      on ChangeValue: SetBit("DB704_MH_Value_Write")
   "DB604_PV_Mixinghead_Mixinghead{0}_Temperature_Connection{2}_PV_Conf_ActV_MaxValueSensor" : Real = PLC DB604_PV_Mixinghead.Mixinghead[0].Temperature_Connection[2].PV_Conf_ActV.MaxValueSensor AT %DB604.DBD382, 1 s
      on ChangeValue: SetBit("DB704_MH_Value_Write")
   "DB604_PV_Mixinghead_Mixinghead{0}_Temperature_Connection{2}_PV_Conf_ActV_MaxSignalResolution" : Real = PLC DB604_PV_Mixinghead.Mixinghead[0].Temperature_Connection[2].PV_Conf_ActV.MaxSignalResolution AT %DB604.DBD386, 1 s
      on ChangeValue: SetBit("DB704_MH_Value_Write")
   "DB604_PV_Mixinghead_Mixinghead{0}_Temperature_Connection{3}_PV_Conf_ActV_ModulNo" : Int = PLC DB604_PV_Mixinghead.Mixinghead[0].Temperature_Connection[3].PV_Conf_ActV.ModulNo AT %DB604.DBW416, 1 s
      on ChangeValue: SetBit("DB704_MH_Value_Write")
   "DB604_PV_Mixinghead_Mixinghead{0}_Temperature_Connection{3}_PV_Conf_ActV_Address" : Int = PLC DB604_PV_Mixinghead.Mixinghead[0].Temperature_Connection[3].PV_Conf_ActV.Address AT %DB604.DBW418, 1 s
      on ChangeValue: SetBit("DB704_MH_Value_Write")
   "DB604_PV_Mixinghead_Mixinghead{0}_Temperature_Connection{3}_PV_Conf_ActV_OffsetSignal" : Int = PLC DB604_PV_Mixinghead.Mixinghead[0].Temperature_Connection[3].PV_Conf_ActV.OffsetSignal AT %DB604.DBW420, 1 s
      on ChangeValue: SetBit("DB704_MH_Value_Write")
   "DB604_PV_Mixinghead_Mixinghead{0}_Temperature_Connection{3}_PV_Conf_ActV_Multiplier" : Real = PLC DB604_PV_Mixinghead.Mixinghead[0].Temperature_Connection[3].PV_Conf_ActV.Multiplier AT %DB604.DBD422, 1 s
      on ChangeValue: SetBit("DB704_MH_Value_Write")
   "DB604_PV_Mixinghead_Mixinghead{0}_Temperature_Connection{3}_PV_Conf_ActV_MinValueSensor" : Real = PLC DB604_PV_Mixinghead.Mixinghead[0].Temperature_Connection[3].PV_Conf_ActV.MinValueSensor AT %DB604.DBD426, 1 s
      on ChangeValue: SetBit("DB704_MH_Value_Write")
   "DB604_PV_Mixinghead_Mixinghead{0}_Temperature_Connection{3}_PV_Conf_ActV_MaxValueSensor" : Real = PLC DB604_PV_Mixinghead.Mixinghead[0].Temperature_Connection[3].PV_Conf_ActV.MaxValueSensor AT %DB604.DBD430, 1 s
      on ChangeValue: SetBit("DB704_MH_Value_Write")
   "DB604_PV_Mixinghead_Mixinghead{0}_Temperature_Connection{3}_PV_Conf_ActV_MaxSignalResolution" : Real = PLC DB604_PV_Mixinghead.Mixinghead[0].Temperature_Connection[3].PV_Conf_ActV.MaxSignalResolution AT %DB604.DBD434, 1 s
      on ChangeValue: SetBit("DB704_MH_Value_Write")
   "DB604_PV_Mixinghead_Mixinghead{0}_Temperature_Connection{4}_PV_Conf_ActV_ModulNo" : Int = PLC DB604_PV_Mixinghead.Mixinghead[0].Temperature_Connection[4].PV_Conf_ActV.ModulNo AT %DB604.DBW464, 1 s
      on ChangeValue: SetBit("DB704_MH_Value_Write")
   "DB604_PV_Mixinghead_Mixinghead{0}_Temperature_Connection{4}_PV_Conf_ActV_Address" : Int = PLC DB604_PV_Mixinghead.Mixinghead[0].Temperature_Connection[4].PV_Conf_ActV.Address AT %DB604.DBW466, 1 s
      on ChangeValue: SetBit("DB704_MH_Value_Write")
   "DB604_PV_Mixinghead_Mixinghead{0}_Temperature_Connection{4}_PV_Conf_ActV_OffsetSignal" : Int = PLC DB604_PV_Mixinghead.Mixinghead[0].Temperature_Connection[4].PV_Conf_ActV.OffsetSignal AT %DB604.DBW468, 1 s
      on ChangeValue: SetBit("DB704_MH_Value_Write")
   "DB604_PV_Mixinghead_Mixinghead{0}_Temperature_Connection{4}_PV_Conf_ActV_Multiplier" : Real = PLC DB604_PV_Mixinghead.Mixinghead[0].Temperature_Connection[4].PV_Conf_ActV.Multiplier AT %DB604.DBD470, 1 s
      on ChangeValue: SetBit("DB704_MH_Value_Write")
   "DB604_PV_Mixinghead_Mixinghead{0}_Temperature_Connection{4}_PV_Conf_ActV_MinValueSensor" : Real = PLC DB604_PV_Mixinghead.Mixinghead[0].Temperature_Connection[4].PV_Conf_ActV.MinValueSensor AT %DB604.DBD474, 1 s
      on ChangeValue: SetBit("DB704_MH_Value_Write")
   "DB604_PV_Mixinghead_Mixinghead{0}_Temperature_Connection{4}_PV_Conf_ActV_MaxValueSensor" : Real = PLC DB604_PV_Mixinghead.Mixinghead[0].Temperature_Connection[4].PV_Conf_ActV.MaxValueSensor AT %DB604.DBD478, 1 s
      on ChangeValue: SetBit("DB704_MH_Value_Write")
   "DB604_PV_Mixinghead_Mixinghead{0}_Temperature_Connection{4}_PV_Conf_ActV_MaxSignalResolution" : Real = PLC DB604_PV_Mixinghead.Mixinghead[0].Temperature_Connection[4].PV_Conf_ActV.MaxSignalResolution AT %DB604.DBD482, 1 s
      on ChangeValue: SetBit("DB704_MH_Value_Write")
   "DB604_PV_Mixinghead_Mixinghead{0}_Temperature_Connection{5}_PV_Conf_ActV_ModulNo" : Int = PLC DB604_PV_Mixinghead.Mixinghead[0].Temperature_Connection[5].PV_Conf_ActV.ModulNo AT %DB604.DBW512, 1 s
      on ChangeValue: SetBit("DB704_MH_Value_Write")
   "DB604_PV_Mixinghead_Mixinghead{0}_Temperature_Connection{5}_PV_Conf_ActV_Address" : Int = PLC DB604_PV_Mixinghead.Mixinghead[0].Temperature_Connection[5].PV_Conf_ActV.Address AT %DB604.DBW514, 1 s
      on ChangeValue: SetBit("DB704_MH_Value_Write")
   "DB604_PV_Mixinghead_Mixinghead{0}_Temperature_Connection{5}_PV_Conf_ActV_OffsetSignal" : Int = PLC DB604_PV_Mixinghead.Mixinghead[0].Temperature_Connection[5].PV_Conf_ActV.OffsetSignal AT %DB604.DBW516, 1 s
      on ChangeValue: SetBit("DB704_MH_Value_Write")
   "DB604_PV_Mixinghead_Mixinghead{0}_Temperature_Connection{5}_PV_Conf_ActV_Multiplier" : Real = PLC DB604_PV_Mixinghead.Mixinghead[0].Temperature_Connection[5].PV_Conf_ActV.Multiplier AT %DB604.DBD518, 1 s
      on ChangeValue: SetBit("DB704_MH_Value_Write")
   "DB604_PV_Mixinghead_Mixinghead{0}_Temperature_Connection{5}_PV_Conf_ActV_MinValueSensor" : Real = PLC DB604_PV_Mixinghead.Mixinghead[0].Temperature_Connection[5].PV_Conf_ActV.MinValueSensor AT %DB604.DBD522, 1 s
      on ChangeValue: SetBit("DB704_MH_Value_Write")
   "DB604_PV_Mixinghead_Mixinghead{0}_Temperature_Connection{5}_PV_Conf_ActV_MaxValueSensor" : Real = PLC DB604_PV_Mixinghead.Mixinghead[0].Temperature_Connection[5].PV_Conf_ActV.MaxValueSensor AT %DB604.DBD526, 1 s
      on ChangeValue: SetBit("DB704_MH_Value_Write")
   "DB604_PV_Mixinghead_Mixinghead{0}_Temperature_Connection{5}_PV_Conf_ActV_MaxSignalResolution" : Real = PLC DB604_PV_Mixinghead.Mixinghead[0].Temperature_Connection[5].PV_Conf_ActV.MaxSignalResolution AT %DB604.DBD530, 1 s
      on ChangeValue: SetBit("DB704_MH_Value_Write")
   "DB604_PV_Mixinghead_Mixinghead{0}_Temperature_Connection{6}_PV_Conf_ActV_ModulNo" : Int = PLC DB604_PV_Mixinghead.Mixinghead[0].Temperature_Connection[6].PV_Conf_ActV.ModulNo AT %DB604.DBW560, 1 s
      on ChangeValue: SetBit("DB704_MH_Value_Write")
   "DB604_PV_Mixinghead_Mixinghead{0}_Temperature_Connection{6}_PV_Conf_ActV_Address" : Int = PLC DB604_PV_Mixinghead.Mixinghead[0].Temperature_Connection[6].PV_Conf_ActV.Address AT %DB604.DBW562, 1 s
      on ChangeValue: SetBit("DB704_MH_Value_Write")
   "DB604_PV_Mixinghead_Mixinghead{0}_Temperature_Connection{6}_PV_Conf_ActV_OffsetSignal" : Int = PLC DB604_PV_Mixinghead.Mixinghead[0].Temperature_Connection[6].PV_Conf_ActV.OffsetSignal AT %DB604.DBW564, 1 s
      on ChangeValue: SetBit("DB704_MH_Value_Write")
   "DB604_PV_Mixinghead_Mixinghead{0}_Temperature_Connection{6}_PV_Conf_ActV_Multiplier" : Real = PLC DB604_PV_Mixinghead.Mixinghead[0].Temperature_Connection[6].PV_Conf_ActV.Multiplier AT %DB604.DBD566, 1 s
      on ChangeValue: SetBit("DB704_MH_Value_Write")
   "DB604_PV_Mixinghead_Mixinghead{0}_Temperature_Connection{6}_PV_Conf_ActV_MinValueSensor" : Real = PLC DB604_PV_Mixinghead.Mixinghead[0].Temperature_Connection[6].PV_Conf_ActV.MinValueSensor AT %DB604.DBD570, 1 s
      on ChangeValue: SetBit("DB704_MH_Value_Write")
   "DB604_PV_Mixinghead_Mixinghead{0}_Temperature_Connection{6}_PV_Conf_ActV_MaxValueSensor" : Real = PLC DB604_PV_Mixinghead.Mixinghead[0].Temperature_Connection[6].PV_Conf_ActV.MaxValueSensor AT %DB604.DBD574, 1 s
      on ChangeValue: SetBit("DB704_MH_Value_Write")
   "DB604_PV_Mixinghead_Mixinghead{0}_Temperature_Connection{6}_PV_Conf_ActV_MaxSignalResolution" : Real = PLC DB604_PV_Mixinghead.Mixinghead[0].Temperature_Connection[6].PV_Conf_ActV.MaxSignalResolution AT %DB604.DBD578, 1 s
      on ChangeValue: SetBit("DB704_MH_Value_Write")
   "DB608_PV_Metering_Metering{0}_MixingRatio_PV_ActV_Value" : Real = PLC DB608_PV_Metering.Metering[0].MixingRatio.PV_ActV.Value AT %DB608.DBD218, 1 s
   "DB608_PV_Metering_HeatexchangerLP{0}_PV_ActV_Value" : Real = PLC DB608_PV_Metering.HeatexchangerLP[0].PV_ActV.Value AT %DB608.DBD3770, 1 s

HMI tags "Last Shot"
   "DB918_ShotResultlast10_FilteredShot{1}_MHNo" : Byte = PLC DB918_ShotResultlast10.FilteredShot[1].MHNo AT %DB918.DBB20, 1 s
   "DB918_ShotResultlast10_FilteredShot{1}_FoamingTime" : Real = PLC DB918_ShotResultlast10.FilteredShot[1].FoamingTime AT %DB918.DBD6, 1 s
   "DB918_ShotResultlast10_FilteredShot{1}_PartWeight" : Real = PLC DB918_ShotResultlast10.FilteredShot[1].PartWeight AT %DB918.DBD10, 1 s
   "DB918_ShotResultlast10_FilteredShot{1}_StationNo" : Byte = PLC DB918_ShotResultlast10.FilteredShot[1].StationNo AT %DB918.DBB18, 1 s
   "DB918_ShotResultlast10_FilteredShot{1}_PartNo" : Int = PLC DB918_ShotResultlast10.FilteredShot[1].PartNo AT %DB918.DBW2, 1 s
   "DB918_ShotResultlast10_FilteredShot{1}_Name{1}" : String[20] = PLC DB918_ShotResultlast10.FilteredShot[1].Name[1] AT %DB918.DBX22.0, 1 s
   "DB918_ShotResultlast10_FilteredShot{1}_Name{2}" : String[20] = PLC DB918_ShotResultlast10.FilteredShot[1].Name[2] AT %DB918.DBX44.0, 1 s
   "DB918_ShotResultlast10_FilteredShot{1}_Flow{1}" : Real = PLC DB918_ShotResultlast10.FilteredShot[1].Flow[1] AT %DB918.DBD154, 1 s
   "DB918_ShotResultlast10_FilteredShot{1}_Flow{2}" : Real = PLC DB918_ShotResultlast10.FilteredShot[1].Flow[2] AT %DB918.DBD158, 1 s
   "DB918_ShotResultlast10_FilteredShot{1}_Pressure{1}" : Real = PLC DB918_ShotResultlast10.FilteredShot[1].Pressure[1] AT %DB918.DBD178, 1 s
   "DB918_ShotResultlast10_FilteredShot{1}_Pressure{2}" : Real = PLC DB918_ShotResultlast10.FilteredShot[1].Pressure[2] AT %DB918.DBD182, 1 s
   "DB918_ShotResultlast10_FilteredShot{1}_Temperature{1}" : Real = PLC DB918_ShotResultlast10.FilteredShot[1].Temperature[1] AT %DB918.DBD202, 1 s
   "DB918_ShotResultlast10_FilteredShot{1}_Temperature{2}" : Real = PLC DB918_ShotResultlast10.FilteredShot[1].Temperature[2] AT %DB918.DBD206, 1 s
   "DB918_ShotResultlast10_FilteredShot{1}_Mixingratio{1}" : Real = PLC DB918_ShotResultlast10.FilteredShot[1].Mixingratio[1] AT %DB918.DBD250, 1 s
   "DB918_ShotResultlast10_FilteredShot{1}_Mixingratio{2}" : Real = PLC DB918_ShotResultlast10.FilteredShot[1].Mixingratio[2] AT %DB918.DBD254, 1 s
   "DB918_ShotResultlast10_FilteredShot{1}_MaterialConsumption{1}" : Real = PLC DB918_ShotResultlast10.FilteredShot[1].MaterialConsumption[1] AT %DB918.DBD226, 1 s
   "DB918_ShotResultlast10_FilteredShot{1}_MaterialConsumption{2}" : Real = PLC DB918_ShotResultlast10.FilteredShot[1].MaterialConsumption[2] AT %DB918.DBD230, 1 s
   "DB918_ShotResultlast10_FilteredShot{2}_PartNo" : Int = PLC DB918_ShotResultlast10.FilteredShot[2].PartNo AT %DB918.DBW288, 1 s
   "DB918_ShotResultlast10_FilteredShot{2}_FoamingTime" : Real = PLC DB918_ShotResultlast10.FilteredShot[2].FoamingTime AT %DB918.DBD292, 1 s
   "DB918_ShotResultlast10_FilteredShot{2}_PartWeight" : Real = PLC DB918_ShotResultlast10.FilteredShot[2].PartWeight AT %DB918.DBD296, 1 s
   "DB918_ShotResultlast10_FilteredShot{2}_StationNo" : Byte = PLC DB918_ShotResultlast10.FilteredShot[2].StationNo AT %DB918.DBB304, 1 s
   "DB918_ShotResultlast10_FilteredShot{2}_MHNo" : Byte = PLC DB918_ShotResultlast10.FilteredShot[2].MHNo AT %DB918.DBB306, 1 s
   "DB918_ShotResultlast10_FilteredShot{2}_Name{1}" : String[20] = PLC DB918_ShotResultlast10.FilteredShot[2].Name[1] AT %DB918.DBX308.0, 1 s
   "DB918_ShotResultlast10_FilteredShot{2}_Name{2}" : String[20] = PLC DB918_ShotResultlast10.FilteredShot[2].Name[2] AT %DB918.DBX330.0, 1 s
   "DB918_ShotResultlast10_FilteredShot{2}_Flow{1}" : Real = PLC DB918_ShotResultlast10.FilteredShot[2].Flow[1] AT %DB918.DBD440, 1 s
   "DB918_ShotResultlast10_FilteredShot{2}_Flow{2}(1)" : Real = PLC DB918_ShotResultlast10.FilteredShot[2].Flow[2] AT %DB918.DBD444, 1 s
   "DB918_ShotResultlast10_FilteredShot{2}_Pressure{1}" : Real = PLC DB918_ShotResultlast10.FilteredShot[2].Pressure[1] AT %DB918.DBD464, 1 s
   "DB918_ShotResultlast10_FilteredShot{2}_Pressure{2}" : Real = PLC DB918_ShotResultlast10.FilteredShot[2].Pressure[2] AT %DB918.DBD468, 1 s
   "DB918_ShotResultlast10_FilteredShot{2}_Temperature{1}" : Real = PLC DB918_ShotResultlast10.FilteredShot[2].Temperature[1] AT %DB918.DBD488, 1 s
   "DB918_ShotResultlast10_FilteredShot{2}_Temperature{2}" : Real = PLC DB918_ShotResultlast10.FilteredShot[2].Temperature[2] AT %DB918.DBD492, 1 s
   "DB918_ShotResultlast10_FilteredShot{2}_MaterialConsumption{1}" : Real = PLC DB918_ShotResultlast10.FilteredShot[2].MaterialConsumption[1] AT %DB918.DBD512, 1 s
   "DB918_ShotResultlast10_FilteredShot{2}_MaterialConsumption{2}" : Real = PLC DB918_ShotResultlast10.FilteredShot[2].MaterialConsumption[2] AT %DB918.DBD516, 1 s
   "DB918_ShotResultlast10_FilteredShot{2}_Mixingratio{1}" : Real = PLC DB918_ShotResultlast10.FilteredShot[2].Mixingratio[1] AT %DB918.DBD536, 1 s
   "DB918_ShotResultlast10_FilteredShot{2}_Mixingratio{2}" : Real = PLC DB918_ShotResultlast10.FilteredShot[2].Mixingratio[2] AT %DB918.DBD540, 1 s
   "DB918_ShotResultlast10_FilteredShot{3}_PartNo" : Int = PLC DB918_ShotResultlast10.FilteredShot[3].PartNo AT %DB918.DBW574, 1 s
   "DB918_ShotResultlast10_FilteredShot{3}_FoamingTime" : Real = PLC DB918_ShotResultlast10.FilteredShot[3].FoamingTime AT %DB918.DBD578, 1 s
   "DB918_ShotResultlast10_FilteredShot{3}_PartWeight" : Real = PLC DB918_ShotResultlast10.FilteredShot[3].PartWeight AT %DB918.DBD582, 1 s
   "DB918_ShotResultlast10_FilteredShot{3}_StationNo" : Byte = PLC DB918_ShotResultlast10.FilteredShot[3].StationNo AT %DB918.DBB590, 1 s
   "DB918_ShotResultlast10_FilteredShot{3}_MHNo" : Byte = PLC DB918_ShotResultlast10.FilteredShot[3].MHNo AT %DB918.DBB592, 1 s
   "DB918_ShotResultlast10_FilteredShot{3}_Name{1}" : String[20] = PLC DB918_ShotResultlast10.FilteredShot[3].Name[1] AT %DB918.DBX594.0, 1 s
   "DB918_ShotResultlast10_FilteredShot{3}_Name{2}" : String[20] = PLC DB918_ShotResultlast10.FilteredShot[3].Name[2] AT %DB918.DBX616.0, 1 s
   "DB918_ShotResultlast10_FilteredShot{3}_Flow{1}" : Real = PLC DB918_ShotResultlast10.FilteredShot[3].Flow[1] AT %DB918.DBD726, 1 s
   "DB918_ShotResultlast10_FilteredShot{3}_Flow{2}" : Real = PLC DB918_ShotResultlast10.FilteredShot[3].Flow[2] AT %DB918.DBD730, 1 s
   "DB918_ShotResultlast10_FilteredShot{3}_Pressure{1}" : Real = PLC DB918_ShotResultlast10.FilteredShot[3].Pressure[1] AT %DB918.DBD750, 1 s
   "DB918_ShotResultlast10_FilteredShot{3}_Pressure{2}" : Real = PLC DB918_ShotResultlast10.FilteredShot[3].Pressure[2] AT %DB918.DBD754, 1 s
   "DB918_ShotResultlast10_FilteredShot{3}_Temperature{1}" : Real = PLC DB918_ShotResultlast10.FilteredShot[3].Temperature[1] AT %DB918.DBD774, 1 s
   "DB918_ShotResultlast10_FilteredShot{3}_Temperature{2}" : Real = PLC DB918_ShotResultlast10.FilteredShot[3].Temperature[2] AT %DB918.DBD778, 1 s
   "DB918_ShotResultlast10_FilteredShot{3}_MaterialConsumption{1}" : Real = PLC DB918_ShotResultlast10.FilteredShot[3].MaterialConsumption[1] AT %DB918.DBD798, 1 s
   "DB918_ShotResultlast10_FilteredShot{3}_MaterialConsumption{2}" : Real = PLC DB918_ShotResultlast10.FilteredShot[3].MaterialConsumption[2] AT %DB918.DBD802, 1 s
   "DB918_ShotResultlast10_FilteredShot{3}_Mixingratio{1}" : Real = PLC DB918_ShotResultlast10.FilteredShot[3].Mixingratio[1] AT %DB918.DBD822, 1 s
   "DB918_ShotResultlast10_FilteredShot{3}_Mixingratio{2}" : Real = PLC DB918_ShotResultlast10.FilteredShot[3].Mixingratio[2] AT %DB918.DBD826, 1 s
   "DB918_ShotResultlast10_FilteredShot{4}_PartNo" : Int = PLC DB918_ShotResultlast10.FilteredShot[4].PartNo AT %DB918.DBW860, 1 s
   "DB918_ShotResultlast10_FilteredShot{4}_FoamingTime" : Real = PLC DB918_ShotResultlast10.FilteredShot[4].FoamingTime AT %DB918.DBD864, 1 s
   "DB918_ShotResultlast10_FilteredShot{4}_PartWeight" : Real = PLC DB918_ShotResultlast10.FilteredShot[4].PartWeight AT %DB918.DBD868, 1 s
   "DB918_ShotResultlast10_FilteredShot{4}_StationNo" : Byte = PLC DB918_ShotResultlast10.FilteredShot[4].StationNo AT %DB918.DBB876, 1 s
   "DB918_ShotResultlast10_FilteredShot{4}_MHNo" : Byte = PLC DB918_ShotResultlast10.FilteredShot[4].MHNo AT %DB918.DBB878, 1 s
   "DB918_ShotResultlast10_FilteredShot{4}_Name{1}" : String[20] = PLC DB918_ShotResultlast10.FilteredShot[4].Name[1] AT %DB918.DBX880.0, 1 s
   "DB918_ShotResultlast10_FilteredShot{4}_Name{2}" : String[20] = PLC DB918_ShotResultlast10.FilteredShot[4].Name[2] AT %DB918.DBX902.0, 1 s
   "DB918_ShotResultlast10_FilteredShot{4}_Flow{1}" : Real = PLC DB918_ShotResultlast10.FilteredShot[4].Flow[1] AT %DB918.DBD1012, 1 s
   "DB918_ShotResultlast10_FilteredShot{4}_Flow{2}" : Real = PLC DB918_ShotResultlast10.FilteredShot[4].Flow[2] AT %DB918.DBD1016, 1 s
   "DB918_ShotResultlast10_FilteredShot{4}_Pressure{1}" : Real = PLC DB918_ShotResultlast10.FilteredShot[4].Pressure[1] AT %DB918.DBD1036, 1 s
   "DB918_ShotResultlast10_FilteredShot{4}_Pressure{2}" : Real = PLC DB918_ShotResultlast10.FilteredShot[4].Pressure[2] AT %DB918.DBD1040, 1 s
   "DB918_ShotResultlast10_FilteredShot{4}_Temperature{1}" : Real = PLC DB918_ShotResultlast10.FilteredShot[4].Temperature[1] AT %DB918.DBD1060, 1 s
   "DB918_ShotResultlast10_FilteredShot{4}_Temperature{2}" : Real = PLC DB918_ShotResultlast10.FilteredShot[4].Temperature[2] AT %DB918.DBD1064, 1 s
   "DB918_ShotResultlast10_FilteredShot{4}_MaterialConsumption{1}" : Real = PLC DB918_ShotResultlast10.FilteredShot[4].MaterialConsumption[1] AT %DB918.DBD1084, 1 s
   "DB918_ShotResultlast10_FilteredShot{4}_MaterialConsumption{2}" : Real = PLC DB918_ShotResultlast10.FilteredShot[4].MaterialConsumption[2] AT %DB918.DBD1088, 1 s
   "DB918_ShotResultlast10_FilteredShot{4}_Mixingratio{1}" : Real = PLC DB918_ShotResultlast10.FilteredShot[4].Mixingratio[1] AT %DB918.DBD1108, 1 s
   "DB918_ShotResultlast10_FilteredShot{4}_Mixingratio{2}" : Real = PLC DB918_ShotResultlast10.FilteredShot[4].Mixingratio[2] AT %DB918.DBD1112, 1 s
   "DB918_ShotResultlast10_FilteredShot{5}_PartNo" : Int = PLC DB918_ShotResultlast10.FilteredShot[5].PartNo AT %DB918.DBW1146, 1 s
   "DB918_ShotResultlast10_FilteredShot{5}_FoamingTime" : Real = PLC DB918_ShotResultlast10.FilteredShot[5].FoamingTime AT %DB918.DBD1150, 1 s
   "DB918_ShotResultlast10_FilteredShot{5}_PartWeight" : Real = PLC DB918_ShotResultlast10.FilteredShot[5].PartWeight AT %DB918.DBD1154, 1 s
   "DB918_ShotResultlast10_FilteredShot{5}_StationNo" : Byte = PLC DB918_ShotResultlast10.FilteredShot[5].StationNo AT %DB918.DBB1162, 1 s
   "DB918_ShotResultlast10_FilteredShot{5}_MHNo" : Byte = PLC DB918_ShotResultlast10.FilteredShot[5].MHNo AT %DB918.DBB1164, 1 s
   "DB918_ShotResultlast10_FilteredShot{5}_Name{1}" : String[20] = PLC DB918_ShotResultlast10.FilteredShot[5].Name[1] AT %DB918.DBX1166.0, 1 s
   "DB918_ShotResultlast10_FilteredShot{5}_Name{2}" : String[20] = PLC DB918_ShotResultlast10.FilteredShot[5].Name[2] AT %DB918.DBX1188.0, 1 s
   "DB918_ShotResultlast10_FilteredShot{5}_Flow{1}" : Real = PLC DB918_ShotResultlast10.FilteredShot[5].Flow[1] AT %DB918.DBD1298, 1 s
   "DB918_ShotResultlast10_FilteredShot{5}_Flow{2}" : Real = PLC DB918_ShotResultlast10.FilteredShot[5].Flow[2] AT %DB918.DBD1302, 1 s
   "DB918_ShotResultlast10_FilteredShot{5}_Pressure{1}" : Real = PLC DB918_ShotResultlast10.FilteredShot[5].Pressure[1] AT %DB918.DBD1322, 1 s
   "DB918_ShotResultlast10_FilteredShot{5}_Pressure{2}" : Real = PLC DB918_ShotResultlast10.FilteredShot[5].Pressure[2] AT %DB918.DBD1326, 1 s
   "DB918_ShotResultlast10_FilteredShot{5}_Temperature{1}" : Real = PLC DB918_ShotResultlast10.FilteredShot[5].Temperature[1] AT %DB918.DBD1346, 1 s
   "DB918_ShotResultlast10_FilteredShot{5}_Temperature{2}" : Real = PLC DB918_ShotResultlast10.FilteredShot[5].Temperature[2] AT %DB918.DBD1350, 1 s
   "DB918_ShotResultlast10_FilteredShot{5}_MaterialConsumption{1}" : Real = PLC DB918_ShotResultlast10.FilteredShot[5].MaterialConsumption[1] AT %DB918.DBD1370, 1 s
   "DB918_ShotResultlast10_FilteredShot{5}_MaterialConsumption{2}" : Real = PLC DB918_ShotResultlast10.FilteredShot[5].MaterialConsumption[2] AT %DB918.DBD1374, 1 s
   "DB918_ShotResultlast10_FilteredShot{5}_Mixingratio{1}" : Real = PLC DB918_ShotResultlast10.FilteredShot[5].Mixingratio[1] AT %DB918.DBD1394, 1 s
   "DB918_ShotResultlast10_FilteredShot{5}_Mixingratio{2}" : Real = PLC DB918_ShotResultlast10.FilteredShot[5].Mixingratio[2] AT %DB918.DBD1398, 1 s
   "DB918_ShotResultlast10_FilteredShot{6}_PartNo" : Int = PLC DB918_ShotResultlast10.FilteredShot[6].PartNo AT %DB918.DBW1432, 1 s
   "DB918_ShotResultlast10_FilteredShot{6}_FoamingTime" : Real = PLC DB918_ShotResultlast10.FilteredShot[6].FoamingTime AT %DB918.DBD1436, 1 s
   "DB918_ShotResultlast10_FilteredShot{6}_PartWeight" : Real = PLC DB918_ShotResultlast10.FilteredShot[6].PartWeight AT %DB918.DBD1440, 1 s
   "DB918_ShotResultlast10_FilteredShot{6}_StationNo" : Byte = PLC DB918_ShotResultlast10.FilteredShot[6].StationNo AT %DB918.DBB1448, 1 s
   "DB918_ShotResultlast10_FilteredShot{6}_MHNo" : Byte = PLC DB918_ShotResultlast10.FilteredShot[6].MHNo AT %DB918.DBB1450, 1 s
   "DB918_ShotResultlast10_FilteredShot{6}_Name{1}" : String[20] = PLC DB918_ShotResultlast10.FilteredShot[6].Name[1] AT %DB918.DBX1452.0, 1 s
   "DB918_ShotResultlast10_FilteredShot{6}_Name{2}" : String[20] = PLC DB918_ShotResultlast10.FilteredShot[6].Name[2] AT %DB918.DBX1474.0, 1 s
   "DB918_ShotResultlast10_FilteredShot{6}_Flow{1}" : Real = PLC DB918_ShotResultlast10.FilteredShot[6].Flow[1] AT %DB918.DBD1584, 1 s
   "DB918_ShotResultlast10_FilteredShot{6}_Flow{2}" : Real = PLC DB918_ShotResultlast10.FilteredShot[6].Flow[2] AT %DB918.DBD1588, 1 s
   "DB918_ShotResultlast10_FilteredShot{6}_Pressure{1}" : Real = PLC DB918_ShotResultlast10.FilteredShot[6].Pressure[1] AT %DB918.DBD1608, 1 s
   "DB918_ShotResultlast10_FilteredShot{6}_Pressure{2}" : Real = PLC DB918_ShotResultlast10.FilteredShot[6].Pressure[2] AT %DB918.DBD1612, 1 s
   "DB918_ShotResultlast10_FilteredShot{6}_Temperature{1}" : Real = PLC DB918_ShotResultlast10.FilteredShot[6].Temperature[1] AT %DB918.DBD1632, 1 s
   "DB918_ShotResultlast10_FilteredShot{6}_Temperature{2}" : Real = PLC DB918_ShotResultlast10.FilteredShot[6].Temperature[2] AT %DB918.DBD1636, 1 s
   "DB918_ShotResultlast10_FilteredShot{6}_MaterialConsumption{1}" : Real = PLC DB918_ShotResultlast10.FilteredShot[6].MaterialConsumption[1] AT %DB918.DBD1656, 1 s
   "DB918_ShotResultlast10_FilteredShot{6}_MaterialConsumption{2}" : Real = PLC DB918_ShotResultlast10.FilteredShot[6].MaterialConsumption[2] AT %DB918.DBD1660, 1 s
   "DB918_ShotResultlast10_FilteredShot{6}_Mixingratio{1}" : Real = PLC DB918_ShotResultlast10.FilteredShot[6].Mixingratio[1] AT %DB918.DBD1680, 1 s
   "DB918_ShotResultlast10_FilteredShot{6}_Mixingratio{2}" : Real = PLC DB918_ShotResultlast10.FilteredShot[6].Mixingratio[2] AT %DB918.DBD1684, 1 s
   "DB918_ShotResultlast10_FilteredShot{1}_PartShotDisableService" : Bool = PLC DB918_ShotResultlast10.FilteredShot[1].PartShotDisableService AT %DB918.DBX286.0, 1 s
   "DB918_ShotResultlast10_FilteredShot{1}_StatusBitManualShot" : Bool = PLC DB918_ShotResultlast10.FilteredShot[1].StatusBitManualShot AT %DB918.DBX286.4, 1 s
   "DB918_ShotResultlast10_FilteredShot{1}_StatusBitAutomaticShot" : Bool = PLC DB918_ShotResultlast10.FilteredShot[1].StatusBitAutomaticShot AT %DB918.DBX286.5, 1 s
   "DB918_ShotResultlast10_FilteredShot{2}_PartShotDisableService" : Bool = PLC DB918_ShotResultlast10.FilteredShot[2].PartShotDisableService AT %DB918.DBX572.0, 1 s
   "DB918_ShotResultlast10_FilteredShot{2}_StatusBitManualShot" : Bool = PLC DB918_ShotResultlast10.FilteredShot[2].StatusBitManualShot AT %DB918.DBX572.4, 1 s
   "DB918_ShotResultlast10_FilteredShot{2}_StatusBitAutomaticShot" : Bool = PLC DB918_ShotResultlast10.FilteredShot[2].StatusBitAutomaticShot AT %DB918.DBX572.5, 1 s
   "DB918_ShotResultlast10_FilteredShot{3}_PartShotDisableService" : Bool = PLC DB918_ShotResultlast10.FilteredShot[3].PartShotDisableService AT %DB918.DBX858.0, 1 s
   "DB918_ShotResultlast10_FilteredShot{3}_StatusBitManualShot" : Bool = PLC DB918_ShotResultlast10.FilteredShot[3].StatusBitManualShot AT %DB918.DBX858.4, 1 s
   "DB918_ShotResultlast10_FilteredShot{3}_StatusBitAutomaticShot" : Bool = PLC DB918_ShotResultlast10.FilteredShot[3].StatusBitAutomaticShot AT %DB918.DBX858.5, 1 s
   "DB918_ShotResultlast10_FilteredShot{4}_PartShotDisableService" : Bool = PLC DB918_ShotResultlast10.FilteredShot[4].PartShotDisableService AT %DB918.DBX1144.0, 1 s
   "DB918_ShotResultlast10_FilteredShot{4}_StatusBitManualShot" : Bool = PLC DB918_ShotResultlast10.FilteredShot[4].StatusBitManualShot AT %DB918.DBX1144.4, 1 s
   "DB918_ShotResultlast10_FilteredShot{4}_StatusBitAutomaticShot" : Bool = PLC DB918_ShotResultlast10.FilteredShot[4].StatusBitAutomaticShot AT %DB918.DBX1144.5, 1 s
   "DB918_ShotResultlast10_FilteredShot{5}_PartShotDisableService" : Bool = PLC DB918_ShotResultlast10.FilteredShot[5].PartShotDisableService AT %DB918.DBX1430.0, 1 s
   "DB918_ShotResultlast10_FilteredShot{5}_StatusBitManualShot" : Bool = PLC DB918_ShotResultlast10.FilteredShot[5].StatusBitManualShot AT %DB918.DBX1430.4, 1 s
   "DB918_ShotResultlast10_FilteredShot{5}_StatusBitAutomaticShot" : Bool = PLC DB918_ShotResultlast10.FilteredShot[5].StatusBitAutomaticShot AT %DB918.DBX1430.5, 1 s
   "DB918_ShotResultlast10_FilteredShot{6}_PartShotDisableService" : Bool = PLC DB918_ShotResultlast10.FilteredShot[6].PartShotDisableService AT %DB918.DBX1716.0, 1 s
   "DB918_ShotResultlast10_FilteredShot{6}_StatusBitManualShot" : Bool = PLC DB918_ShotResultlast10.FilteredShot[6].StatusBitManualShot AT %DB918.DBX1716.4, 1 s
   "DB918_ShotResultlast10_FilteredShot{6}_StatusBitAutomaticShot" : Bool = PLC DB918_ShotResultlast10.FilteredShot[6].StatusBitAutomaticShot AT %DB918.DBX1716.5, 1 s

HMI tags "General View"
   "DB602_PV_Tank_Tank{1}_Temp_PV_ActV_Value" : Real = PLC DB602_PV_Tank.Tank[1].Temp.PV_ActV.Value AT %DB602.DBD266, 1 s
   "DB602_PV_Tank_Tank{1}_Level_PV_ActV_Value" : Real = PLC DB602_PV_Tank.Tank[1].Level.PV_ActV.Value AT %DB602.DBD314, 1 s
   "DB602_PV_Tank_Tank{2}_Level_PV_ActV_Value" : Real = PLC DB602_PV_Tank.Tank[2].Level.PV_ActV.Value AT %DB602.DBD554, 1 s
   "DB602_PV_Tank_Tank{2}_Temp_PV_ActV_Value" : Real = PLC DB602_PV_Tank.Tank[2].Temp.PV_ActV.Value AT %DB602.DBD506, 1 s
   "DB608_PV_Metering_Metering{1}_Flow_PV_ActV_Value" : Real = PLC DB608_PV_Metering.Metering[1].Flow.PV_ActV.Value AT %DB608.DBD266, 1 s
   "DB608_PV_Metering_Metering{1}_Pressure_PV_ActV_Value" : Real = PLC DB608_PV_Metering.Metering[1].Pressure.PV_ActV.Value AT %DB608.DBD314, 1 s
   "DB608_PV_Metering_Metering{1}_MixingRatio_PV_ActV_Value" : Real = PLC DB608_PV_Metering.Metering[1].MixingRatio.PV_ActV.Value AT %DB608.DBD458, 1 s
   "DB608_PV_Metering_Metering{2}_Flow_PV_ActV_Value" : Real = PLC DB608_PV_Metering.Metering[2].Flow.PV_ActV.Value AT %DB608.DBD506, 1 s
   "DB608_PV_Metering_Metering{2}_Pressure_PV_ActV_Value" : Real = PLC DB608_PV_Metering.Metering[2].Pressure.PV_ActV.Value AT %DB608.DBD554, 1 s
   "DB608_PV_Metering_Metering{2}_MixingRatio_PV_ActV_Value" : Real = PLC DB608_PV_Metering.Metering[2].MixingRatio.PV_ActV.Value AT %DB608.DBD698, 1 s
   "DB619_State_MPart_ActMHPressureMa{1}_Comp{1}" : Real = PLC DB619_State_MPart.ActMHPressureMa[1].Comp[1] AT %DB619.DBD2480, 1 s
   "DB619_State_MPart_ActMHPressureMa{1}_Comp{2}" : Real = PLC DB619_State_MPart.ActMHPressureMa[1].Comp[2] AT %DB619.DBD2484, 1 s
   "DB619_State_MPart_ActMHTemperatureMa{1}_Comp{1}" : Real = PLC DB619_State_MPart.ActMHTemperatureMa[1].Comp[1] AT %DB619.DBD2720, 1 s
   "DB619_State_MPart_ActMHTemperatureMa{1}_Comp{2}" : Real = PLC DB619_State_MPart.ActMHTemperatureMa[1].Comp[2] AT %DB619.DBD2724, 1 s
   "DB619_State_MPart_ActMHInerting{1}_Total_Flow_N2_Visu" : Real = PLC DB619_State_MPart.ActMHInerting[1].Total_Flow_N2_Visu AT %DB619.DBD3326, 1 s

